(* Logix 5000 project; controller PLC_MCC1300_75F1 vendor 1 type 14 code 166 rev 32.11; software revision 32.04; part 58 of 83 *)
(* tags used below, declared in another part *)
   CM_AreaStackerToLine_JS1_Sync : CM_AreaStackerToLine;
   CM_ConveyorStackerToLine_JS1_Sync : CM_ConveyorStackerToLine;
   CM_DATA_Z410_Rx_Sync : UDT_PlateData_Convoy;
   CM_LineToConveyorStacker_JS1 : CM_LineToConveyorStacker;
   GP_AccessArea_M311S_STC : GP_AccessArea_STC;
   GP_ConvertDataFromStacker : GP_ConvertDataFromStacker;
   Gp_SpaceConvUtilities_V1 : GP_SpaceConvUtilities_V1;
   M311 : MAC_Conveyor;
   M311_SpaceConv_Utilities : SpaceConv_Utilities;
   M312 : MAC_Conveyor_Single;
   M312_ALM : MAC_Conveyor_ALM;
   M312_Data : UDT_Convoy_SL;
   M312_dTractionRecovery_M3 : DINT;
   M312_dTractionRecovery_M4 : DINT;
   M312_HMR : MAC_Conveyor_HMR;
   M312_HMW : MAC_Conveyor_HMW;
   M312_M3_DR_IN_MAM : MOTION_INSTRUCTION;
   M312_M3_DR_IN_MRP : MOTION_INSTRUCTION;
   M312_SpaceConv_Utilities : SpaceConv_Utilities;
   M312_TON_FrontSquarLeft_timeout : TIMER;
   M312_TON_FrontSquarRight_timeout : TIMER;
   M312_TON_LatSquarLeft_timeout : TIMER;
   M312_TON_LatSquarRight_timeout : TIMER;
   M312_TON_Synchro_timeout : TIMER;
   M312_xEnableTractionRecovering : BOOL;
   M312_xFrontLeftTimeout : BOOL;
   M312_xFrontRightTimeout : BOOL;
   M312_xLateralTractionRecovered : BOOL;
   M312_xLatLeftTimeout : BOOL;
   M312_xLatRightTimeout : BOOL;
   M312_xSendCulletReqActive : BOOL;
   M312_xSensorTimeout : BOOL;
   O : INT[128];
   TMP_CenterLites : BOOL;
   TMP_d : DINT;
   TMP_DistanceLateralSquaringToCenter : DINT;
   TMP_dOffsetLoadUnload_cmm : DINT;
   TMP_SendToCullet : BOOL;
   TMP_xConveyorOfStartCleaning : BOOL;
   TMP_xEnableZoneCleaning : BOOL;
   TMP_xLiteThisDestPresent : BOOL;
   xAlwaysON : BOOL;
   Z401 : MAC_Zone;
   Z401S_INPUT_xSafetyAreaPopup : BOOL;
(* MainProgram, continued *)

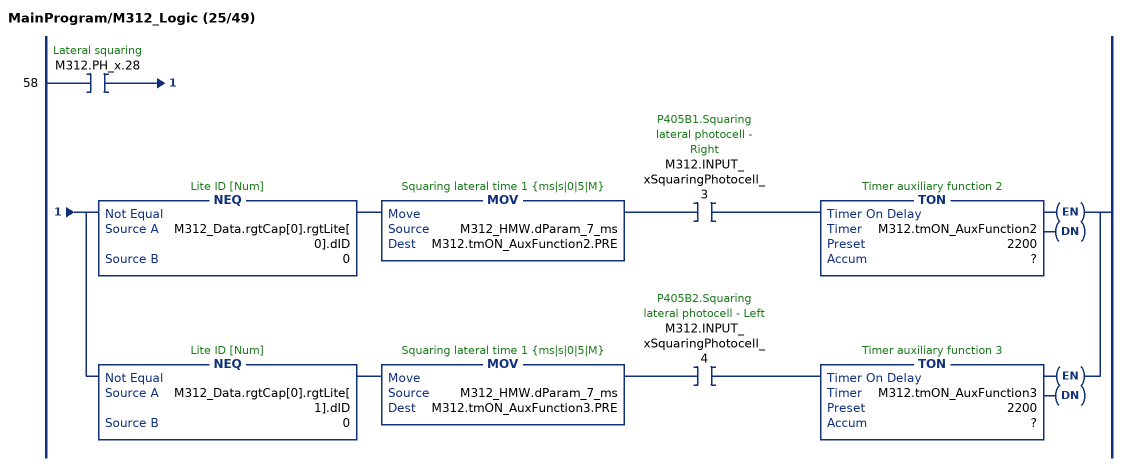
   [picture p958: MainProgram/M312_Logic rungs 58-58]
   58: XIC(M312.PH_x.28)[NEQ(M312_Data.rgtCap[0].rgtLite[0].dID,0) MOV(M312_HMW.dParam_7_ms,M312.tmON_AuxFunction2.PRE) XIC(M312.INPUT_xSquaringPhotocell_3) TON(M312.tmON_AuxFunction2,?,?) ,NEQ(M312_Data.rgtCap[0].rgtLite[1].dID,0) MOV(M312_HMW.dParam_7_ms,M312.tmON_AuxFunction3.PRE) XIC(M312.INPUT_xSquaringPhotocell_4) TON(M312.tmON_AuxFunction3,?,?) ];
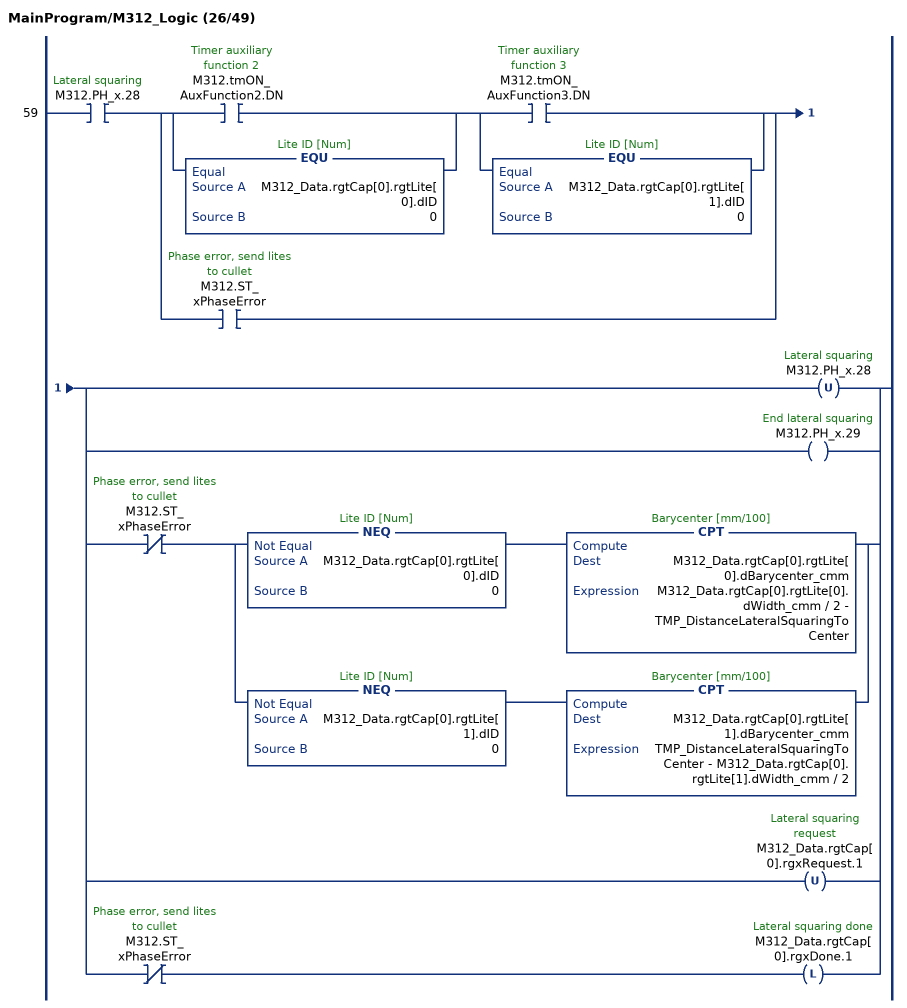
   59: XIC(M312.PH_x.28)[[XIC(M312.tmON_AuxFunction2.DN) ,EQU(M312_Data.rgtCap[0].rgtLite[0].dID,0) ] [XIC(M312.tmON_AuxFunction3.DN) ,EQU(M312_Data.rgtCap[0].rgtLite[1].dID,0) ] ,XIC(M312.ST_xPhaseError) ][OTU(M312.PH_x.28) ,OTE(M312.PH_x.29) ,XIO(M312.ST_xPhaseError) [NEQ(M312_Data.rgtCap[0].rgtLite[0].dID,0) CPT(M312_Data.rgtCap[0].rgtLite[0].dBarycenter_cmm,M312_Data.rgtCap[0].rgtLite[0].dWidth_cmm / 2 - TMP_DistanceLateralSquaringToCenter) ,NEQ(M312_Data.rgtCap[0].rgtLite[1].dID,0) CPT(M312_Data.rgtCap[0].rgtLite[1].dBarycenter_cmm,TMP_DistanceLateralSquaringToCenter - M312_Data.rgtCap[0].rgtLite[1].dWidth_cmm / 2) ] ,OTU(M312_Data.rgtCap[0].rgxRequest.1) ,XIO(M312.ST_xPhaseError) OTL(M312_Data.rgtCap[0].rgxDone.1) ];
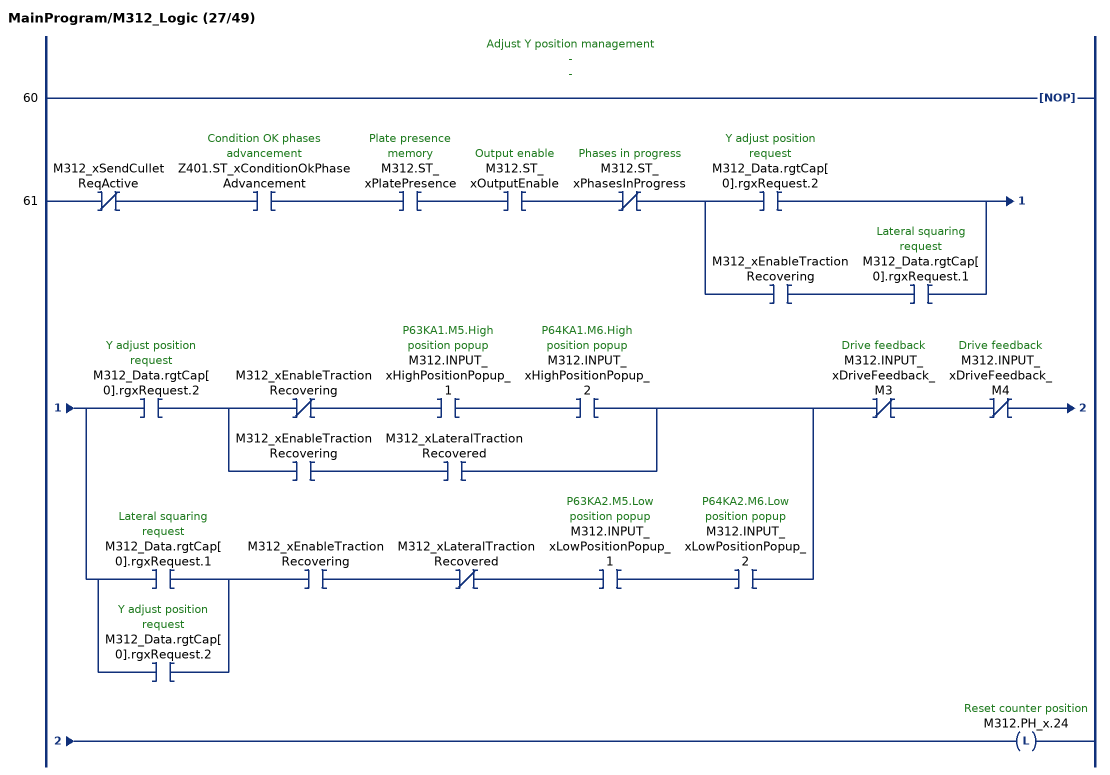
   // Adjust Y position management
   // -
   // -
   60: NOP();
   61: XIO(M312_xSendCulletReqActive)XIC(Z401.ST_xConditionOkPhaseAdvancement)XIC(M312.ST_xPlatePresence)XIC(M312.ST_xOutputEnable)XIO(M312.ST_xPhasesInProgress)[XIC(M312_Data.rgtCap[0].rgxRequest.2) ,XIC(M312_xEnableTractionRecovering) XIC(M312_Data.rgtCap[0].rgxRequest.1) ][XIC(M312_Data.rgtCap[0].rgxRequest.2) [XIO(M312_xEnableTractionRecovering) XIC(M312.INPUT_xHighPositionPopup_1) XIC(M312.INPUT_xHighPositionPopup_2) ,XIC(M312_xEnableTractionRecovering) XIC(M312_xLateralTractionRecovered) ] ,[XIC(M312_Data.rgtCap[0].rgxRequest.1) ,XIC(M312_Data.rgtCap[0].rgxRequest.2) ] XIC(M312_xEnableTractionRecovering) XIO(M312_xLateralTractionRecovered) XIC(M312.INPUT_xLowPositionPopup_1) XIC(M312.INPUT_xLowPositionPopup_2) ]XIO(M312.INPUT_xDriveFeedback_M3)XIO(M312.INPUT_xDriveFeedback_M4)OTL(M312.PH_x.24);
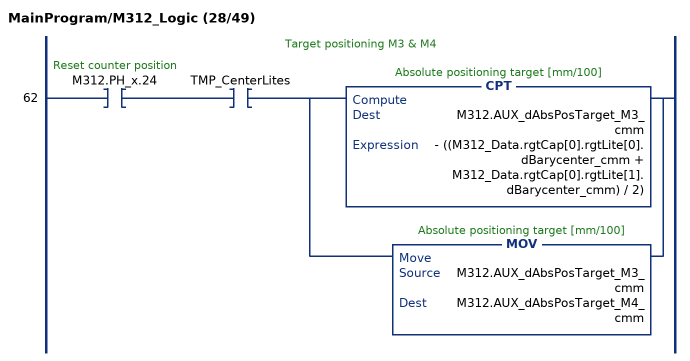
   // Target positioning M3 & M4
   62: XIC(M312.PH_x.24)XIC(TMP_CenterLites)[CPT(M312.AUX_dAbsPosTarget_M3_cmm,- ((M312_Data.rgtCap[0].rgtLite[0].dBarycenter_cmm + M312_Data.rgtCap[0].rgtLite[1].dBarycenter_cmm) / 2)) ,MOV(M312.AUX_dAbsPosTarget_M3_cmm,M312.AUX_dAbsPosTarget_M4_cmm) ];
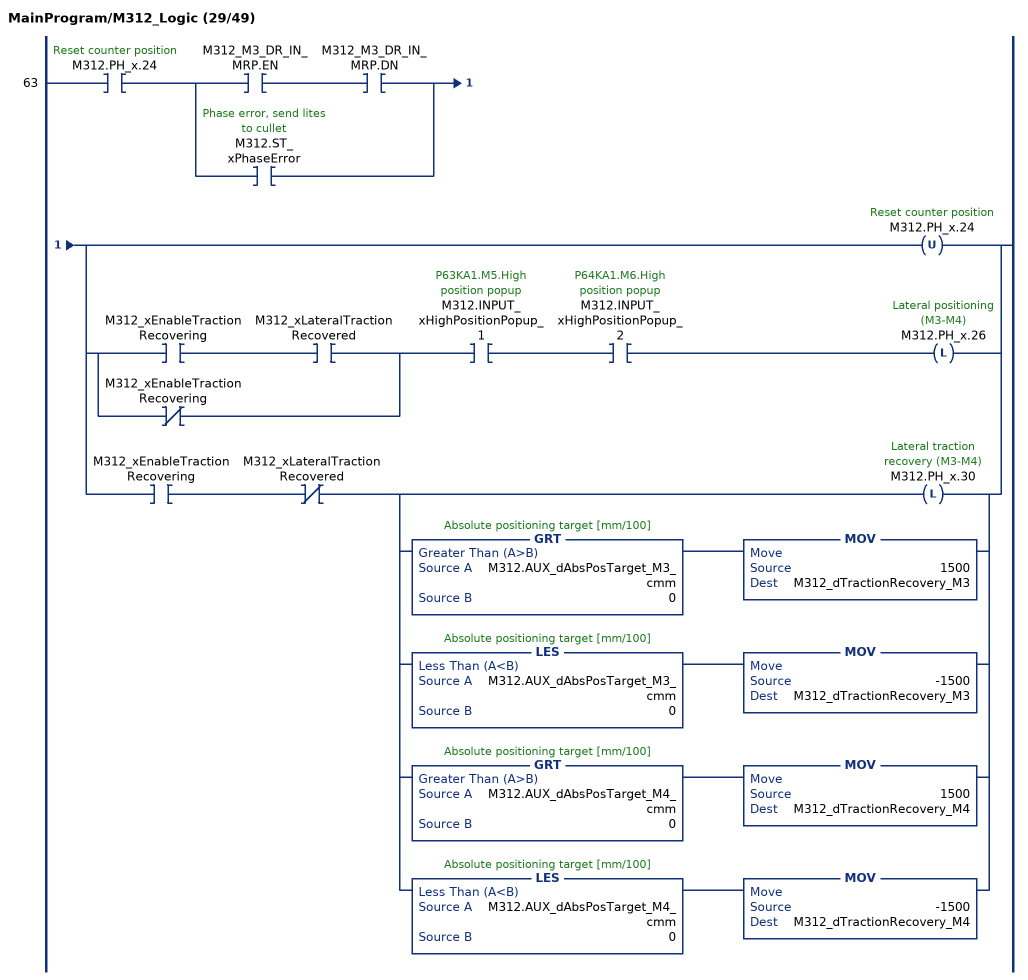
   63: XIC(M312.PH_x.24)[XIC(M312_M3_DR_IN_MRP.EN) XIC(M312_M3_DR_IN_MRP.DN) ,XIC(M312.ST_xPhaseError) ][OTU(M312.PH_x.24) ,[XIC(M312_xEnableTractionRecovering) XIC(M312_xLateralTractionRecovered) ,XIO(M312_xEnableTractionRecovering) ] XIC(M312.INPUT_xHighPositionPopup_1) XIC(M312.INPUT_xHighPositionPopup_2) OTL(M312.PH_x.26) ,XIC(M312_xEnableTractionRecovering) XIO(M312_xLateralTractionRecovered) [OTL(M312.PH_x.30) ,[GRT(M312.AUX_dAbsPosTarget_M3_cmm,0) MOV(1500,M312_dTractionRecovery_M3) ,LES(M312.AUX_dAbsPosTarget_M3_cmm,0) MOV(-1500,M312_dTractionRecovery_M3) ,GRT(M312.AUX_dAbsPosTarget_M4_cmm,0) MOV(1500,M312_dTractionRecovery_M4) ,LES(M312.AUX_dAbsPosTarget_M4_cmm,0) MOV(-1500,M312_dTractionRecovery_M4) ] ] ];
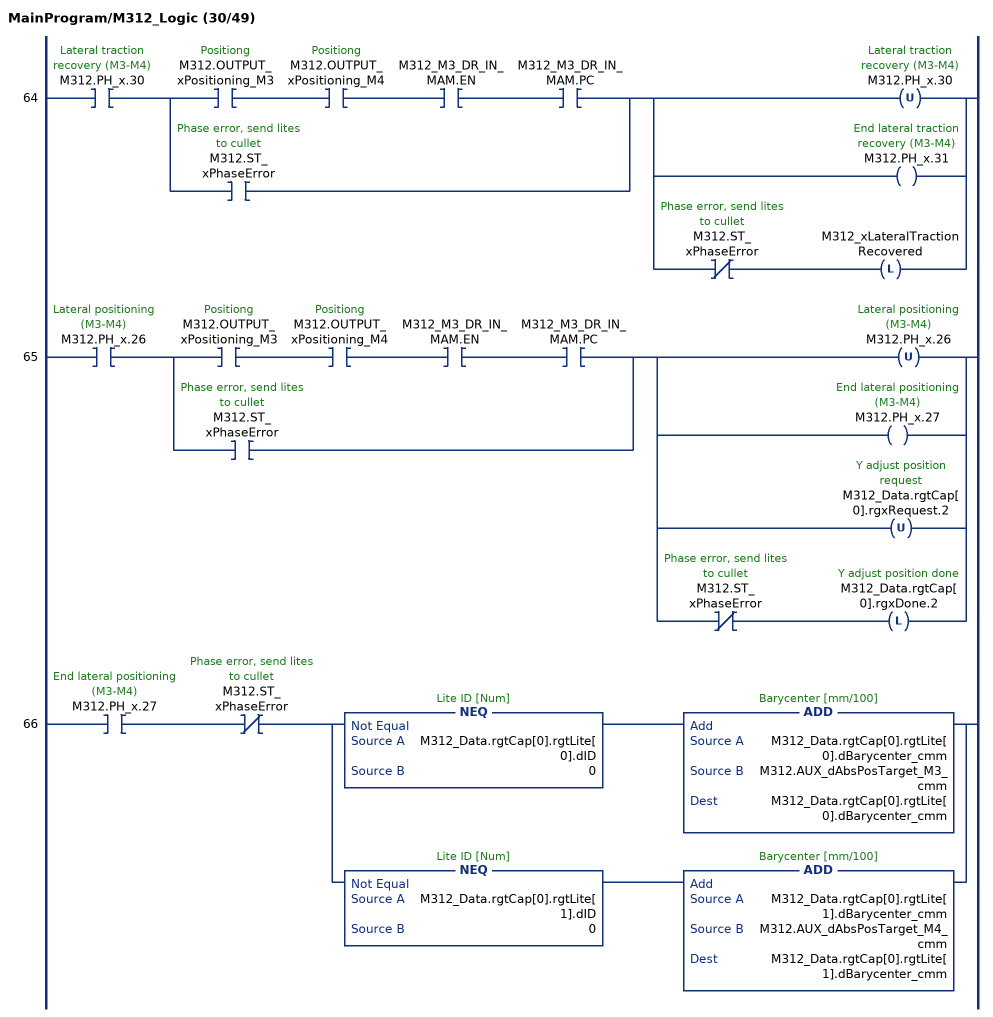
   64: XIC(M312.PH_x.30)[XIC(M312.OUTPUT_xPositioning_M3) XIC(M312.OUTPUT_xPositioning_M4) XIC(M312_M3_DR_IN_MAM.EN) XIC(M312_M3_DR_IN_MAM.PC) ,XIC(M312.ST_xPhaseError) ][OTU(M312.PH_x.30) ,OTE(M312.PH_x.31) ,XIO(M312.ST_xPhaseError) OTL(M312_xLateralTractionRecovered) ];
   65: XIC(M312.PH_x.26)[XIC(M312.OUTPUT_xPositioning_M3) XIC(M312.OUTPUT_xPositioning_M4) XIC(M312_M3_DR_IN_MAM.EN) XIC(M312_M3_DR_IN_MAM.PC) ,XIC(M312.ST_xPhaseError) ][OTU(M312.PH_x.26) ,OTE(M312.PH_x.27) ,OTU(M312_Data.rgtCap[0].rgxRequest.2) ,XIO(M312.ST_xPhaseError) OTL(M312_Data.rgtCap[0].rgxDone.2) ];
   66: XIC(M312.PH_x.27)XIO(M312.ST_xPhaseError)[NEQ(M312_Data.rgtCap[0].rgtLite[0].dID,0) ADD(M312_Data.rgtCap[0].rgtLite[0].dBarycenter_cmm,M312.AUX_dAbsPosTarget_M3_cmm,M312_Data.rgtCap[0].rgtLite[0].dBarycenter_cmm) ,NEQ(M312_Data.rgtCap[0].rgtLite[1].dID,0) ADD(M312_Data.rgtCap[0].rgtLite[1].dBarycenter_cmm,M312.AUX_dAbsPosTarget_M4_cmm,M312_Data.rgtCap[0].rgtLite[1].dBarycenter_cmm) ];
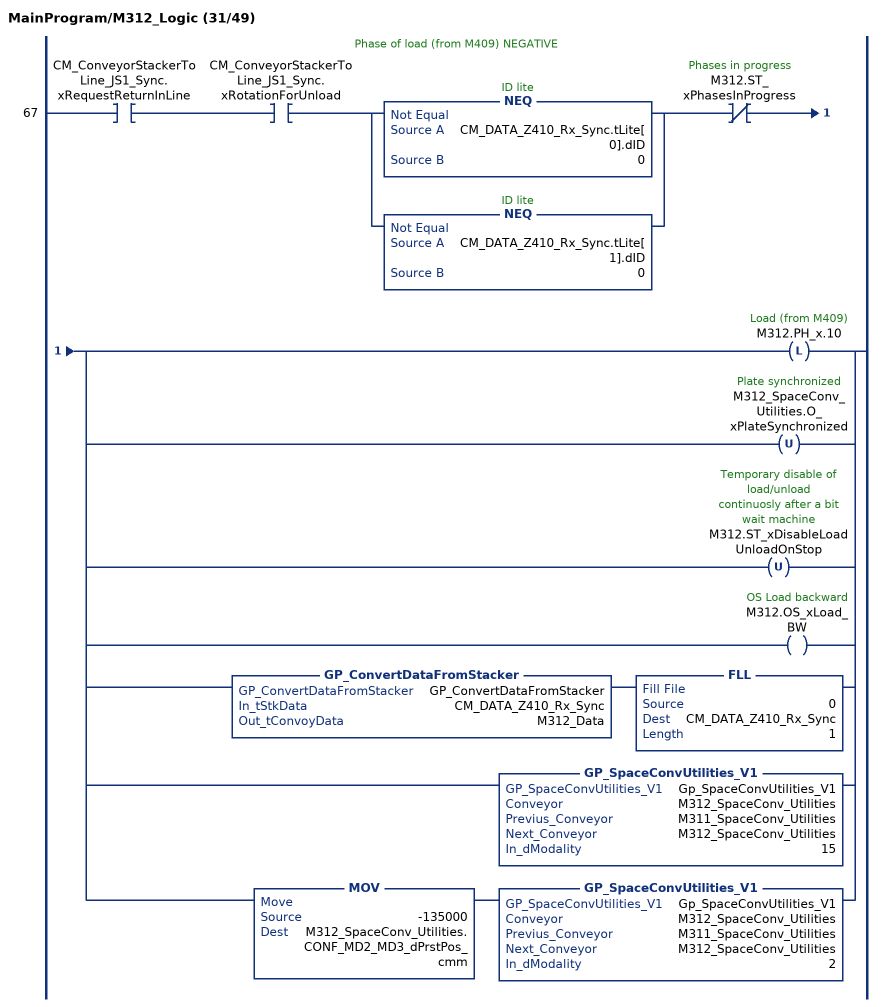
   // Phase of load (from M409) NEGATIVE
   67: XIC(CM_ConveyorStackerToLine_JS1_Sync.xRequestReturnInLine)XIC(CM_ConveyorStackerToLine_JS1_Sync.xRotationForUnload)[NEQ(CM_DATA_Z410_Rx_Sync.tLite[0].dID,0) ,NEQ(CM_DATA_Z410_Rx_Sync.tLite[1].dID,0) ]XIO(M312.ST_xPhasesInProgress)[OTL(M312.PH_x.10) ,OTU(M312_SpaceConv_Utilities.O_xPlateSynchronized) ,OTU(M312.ST_xDisableLoadUnloadOnStop) ,OTE(M312.OS_xLoad_BW) ,GP_ConvertDataFromStacker(GP_ConvertDataFromStacker,CM_DATA_Z410_Rx_Sync,M312_Data) FLL(0,CM_DATA_Z410_Rx_Sync,1) ,GP_SpaceConvUtilities_V1(Gp_SpaceConvUtilities_V1,M312_SpaceConv_Utilities,M311_SpaceConv_Utilities,M312_SpaceConv_Utilities,15) ,MOV(-135000,M312_SpaceConv_Utilities.CONF_MD2_MD3_dPrstPos_cmm) GP_SpaceConvUtilities_V1(Gp_SpaceConvUtilities_V1,M312_SpaceConv_Utilities,M311_SpaceConv_Utilities,M312_SpaceConv_Utilities,2) ];
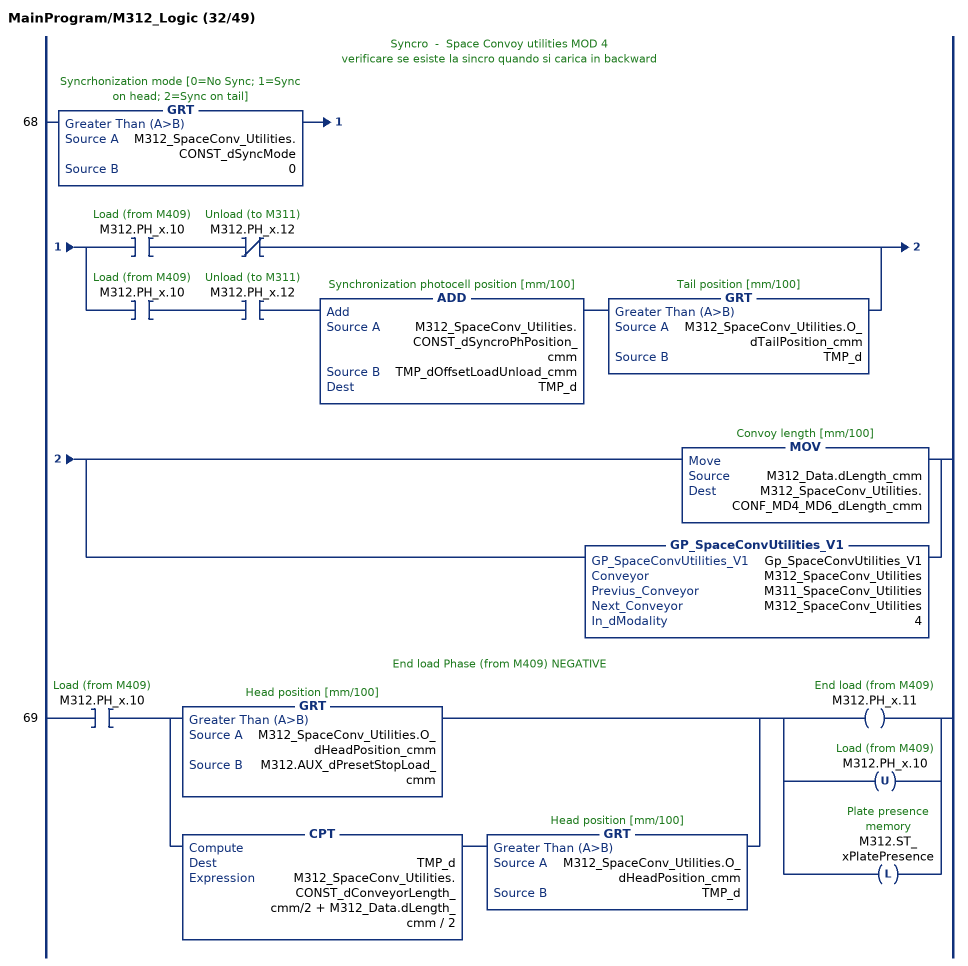
   // Syncro  -  Space Convoy utilities MOD 4
   // verificare se esiste la sincro quando si carica in backward
   68: GRT(M312_SpaceConv_Utilities.CONST_dSyncMode,0)[XIC(M312.PH_x.10) XIO(M312.PH_x.12) ,XIC(M312.PH_x.10) XIC(M312.PH_x.12) ADD(M312_SpaceConv_Utilities.CONST_dSyncroPhPosition_cmm,TMP_dOffsetLoadUnload_cmm,TMP_d) GRT(M312_SpaceConv_Utilities.O_dTailPosition_cmm,TMP_d) ][MOV(M312_Data.dLength_cmm,M312_SpaceConv_Utilities.CONF_MD4_MD6_dLength_cmm) ,GP_SpaceConvUtilities_V1(Gp_SpaceConvUtilities_V1,M312_SpaceConv_Utilities,M311_SpaceConv_Utilities,M312_SpaceConv_Utilities,4) ];
   // End load Phase (from M409) NEGATIVE
   69: XIC(M312.PH_x.10)[GRT(M312_SpaceConv_Utilities.O_dHeadPosition_cmm,M312.AUX_dPresetStopLoad_cmm) ,CPT(TMP_d,M312_SpaceConv_Utilities.CONST_dConveyorLength_cmm/2 + M312_Data.dLength_cmm / 2) GRT(M312_SpaceConv_Utilities.O_dHeadPosition_cmm,TMP_d) ][OTE(M312.PH_x.11) ,OTU(M312.PH_x.10) ,OTL(M312.ST_xPlatePresence) ];
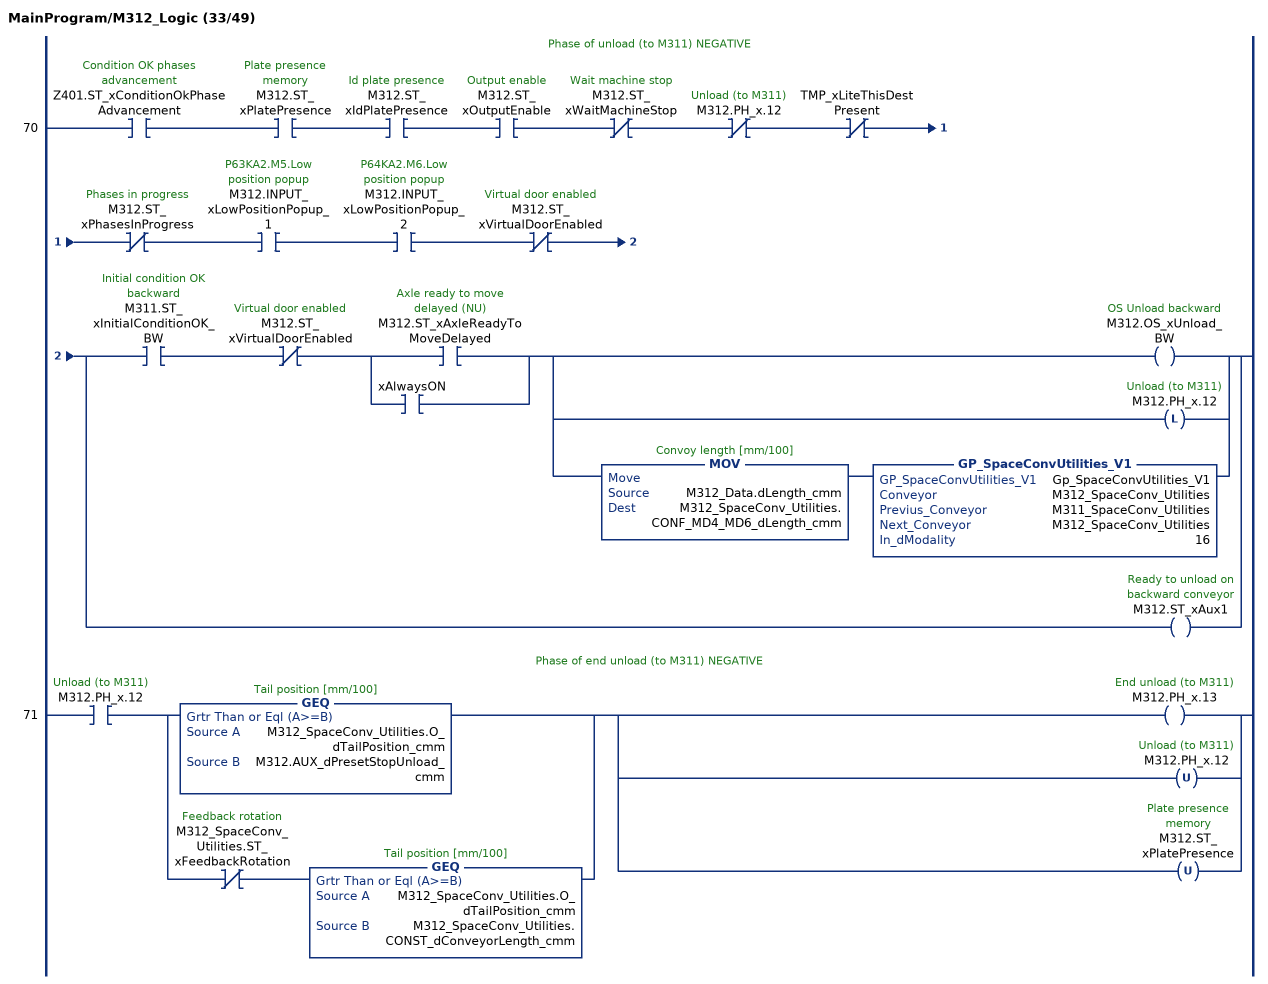
   // Phase of unload (to M311) NEGATIVE
   70: XIC(Z401.ST_xConditionOkPhaseAdvancement)XIC(M312.ST_xPlatePresence)XIC(M312.ST_xIdPlatePresence)XIC(M312.ST_xOutputEnable)XIO(M312.ST_xWaitMachineStop)XIO(M312.PH_x.12)XIO(TMP_xLiteThisDestPresent)XIO(M312.ST_xPhasesInProgress)XIC(M312.INPUT_xLowPositionPopup_1)XIC(M312.INPUT_xLowPositionPopup_2)XIO(M312.ST_xVirtualDoorEnabled)[XIC(M311.ST_xInitialConditionOK_BW) XIO(M312.ST_xVirtualDoorEnabled) [XIC(M312.ST_xAxleReadyToMoveDelayed) ,XIC(xAlwaysON) ] [OTE(M312.OS_xUnload_BW) ,OTL(M312.PH_x.12) ,MOV(M312_Data.dLength_cmm,M312_SpaceConv_Utilities.CONF_MD4_MD6_dLength_cmm) GP_SpaceConvUtilities_V1(Gp_SpaceConvUtilities_V1,M312_SpaceConv_Utilities,M311_SpaceConv_Utilities,M312_SpaceConv_Utilities,16) ] ,OTE(M312.ST_xAux1) ];
   // Phase of end unload (to M311) NEGATIVE
   71: XIC(M312.PH_x.12)[GEQ(M312_SpaceConv_Utilities.O_dTailPosition_cmm,M312.AUX_dPresetStopUnload_cmm) ,XIO(M312_SpaceConv_Utilities.ST_xFeedbackRotation) GEQ(M312_SpaceConv_Utilities.O_dTailPosition_cmm,M312_SpaceConv_Utilities.CONST_dConveyorLength_cmm) ][OTE(M312.PH_x.13) ,OTU(M312.PH_x.12) ,OTU(M312.ST_xPlatePresence) ];